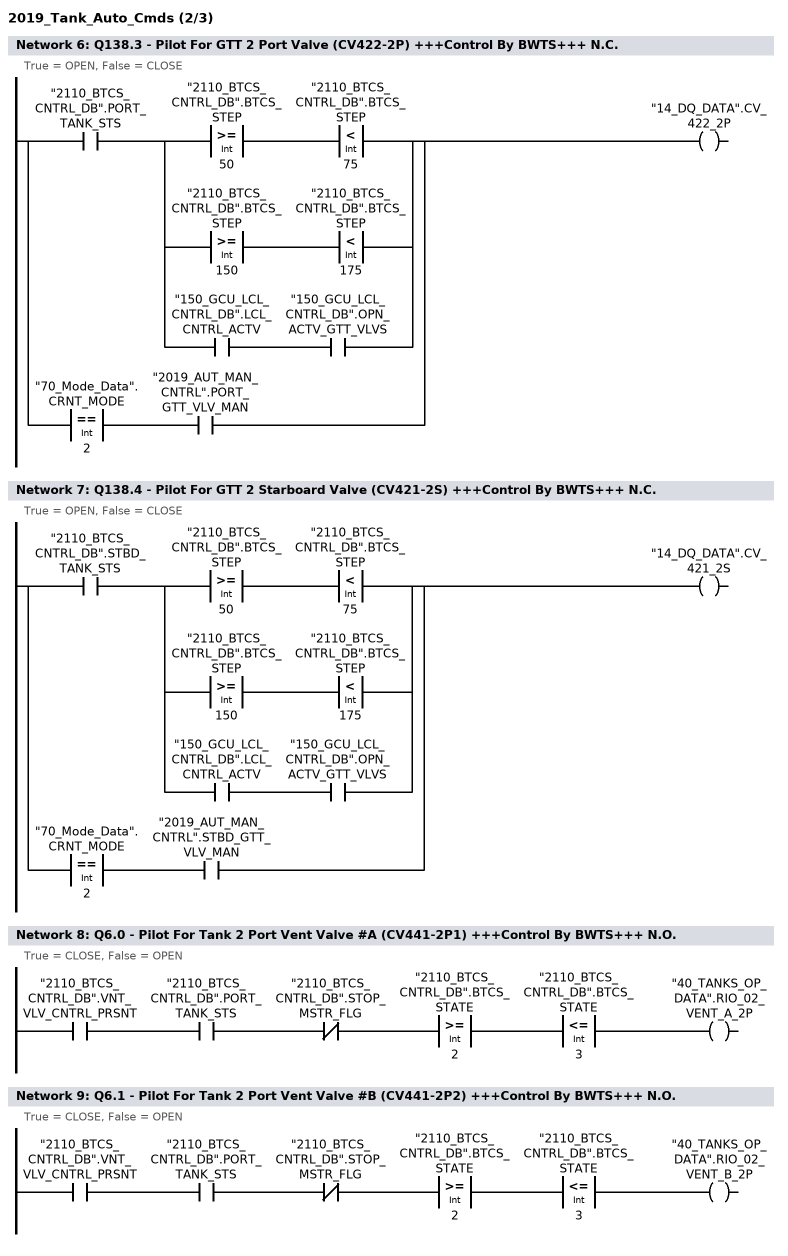
   RUNG wire#powerrail
      Contact( "2110_BTCS_CNTRL_DB".PORT_TANK_STS )
      wire#w1
      { S7_Templates := "SrcType := Int" } GE_Contact(in1 := "2110_BTCS_CNTRL_DB".BTCS_STEP, in2 := 50)
      { S7_Templates := "SrcType := Int" } LT_Contact(in1 := "2110_BTCS_CNTRL_DB".BTCS_STEP, in2 := 75)
      wire#w2
      Coil( "14_DQ_DATA".CV_422_2P )
   END_RUNG
   RUNG wire#w1
      { S7_Templates := "SrcType := Int" } GE_Contact(in1 := "2110_BTCS_CNTRL_DB".BTCS_STEP, in2 := 150)
      { S7_Templates := "SrcType := Int" } LT_Contact(in1 := "2110_BTCS_CNTRL_DB".BTCS_STEP, in2 := 175)
   END_RUNG wire#w2
   RUNG wire#w1
      Contact( "150_GCU_LCL_CNTRL_DB".LCL_CNTRL_ACTV )
      Contact( "150_GCU_LCL_CNTRL_DB".OPN_ACTV_GTT_VLVS )
   END_RUNG wire#w2
   RUNG wire#powerrail
      { S7_Templates := "SrcType := Int" } EQ_Contact(in1 := "70_Mode_Data".CRNT_MODE, in2 := 2)
      Contact( "2019_AUT_MAN_CNTRL".PORT_GTT_VLV_MAN )
   END_RUNG wire#w2
   // the same network as SCL:
   "14_DQ_DATA".CV_422_2P := ("2110_BTCS_CNTRL_DB".PORT_TANK_STS AND ((("2110_BTCS_CNTRL_DB".BTCS_STEP >= 50) AND ("2110_BTCS_CNTRL_DB".BTCS_STEP < 75)) OR (("2110_BTCS_CNTRL_DB".BTCS_STEP >= 150) AND ("2110_BTCS_CNTRL_DB".BTCS_STEP < 175)) OR ("150_GCU_LCL_CNTRL_DB".LCL_CNTRL_ACTV AND "150_GCU_LCL_CNTRL_DB".OPN_ACTV_GTT_VLVS))) OR (("70_Mode_Data".CRNT_MODE = 2) AND "2019_AUT_MAN_CNTRL".PORT_GTT_VLV_MAN);
END_REGION

REGION Network 7: Q138.4 - Pilot For GTT 2 Starboard Valve (CV421-2S) +++Control By BWTS+++ N.C.
   // True = OPEN, False = CLOSE
   RUNG wire#powerrail
      Contact( "2110_BTCS_CNTRL_DB".STBD_TANK_STS )
      wire#w1
      { S7_Templates := "SrcType := Int" } GE_Contact(in1 := "2110_BTCS_CNTRL_DB".BTCS_STEP, in2 := 50)
      { S7_Templates := "SrcType := Int" } LT_Contact(in1 := "2110_BTCS_CNTRL_DB".BTCS_STEP, in2 := 75)
      wire#w2
      Coil( "14_DQ_DATA".CV_421_2S )
   END_RUNG
   RUNG wire#w1
      { S7_Templates := "SrcType := Int" } GE_Contact(in1 := "2110_BTCS_CNTRL_DB".BTCS_STEP, in2 := 150)
      { S7_Templates := "SrcType := Int" } LT_Contact(in1 := "2110_BTCS_CNTRL_DB".BTCS_STEP, in2 := 175)
   END_RUNG wire#w2
   RUNG wire#w1
      Contact( "150_GCU_LCL_CNTRL_DB".LCL_CNTRL_ACTV )
      Contact( "150_GCU_LCL_CNTRL_DB".OPN_ACTV_GTT_VLVS )
   END_RUNG wire#w2
   RUNG wire#powerrail
      { S7_Templates := "SrcType := Int" } EQ_Contact(in1 := "70_Mode_Data".CRNT_MODE, in2 := 2)
      Contact( "2019_AUT_MAN_CNTRL".STBD_GTT_VLV_MAN )
   END_RUNG wire#w2
   // the same network as SCL:
   "14_DQ_DATA".CV_421_2S := ("2110_BTCS_CNTRL_DB".STBD_TANK_STS AND ((("2110_BTCS_CNTRL_DB".BTCS_STEP >= 50) AND ("2110_BTCS_CNTRL_DB".BTCS_STEP < 75)) OR (("2110_BTCS_CNTRL_DB".BTCS_STEP >= 150) AND ("2110_BTCS_CNTRL_DB".BTCS_STEP < 175)) OR ("150_GCU_LCL_CNTRL_DB".LCL_CNTRL_ACTV AND "150_GCU_LCL_CNTRL_DB".OPN_ACTV_GTT_VLVS))) OR (("70_Mode_Data".CRNT_MODE = 2) AND "2019_AUT_MAN_CNTRL".STBD_GTT_VLV_MAN);
END_REGION

REGION Network 8: Q6.0 - Pilot For Tank 2 Port Vent Valve #A (CV441-2P1) +++Control By BWTS+++ N.O.
   // True = CLOSE, False = OPEN
   RUNG wire#powerrail
      Contact( "2110_BTCS_CNTRL_DB".VNT_VLV_CNTRL_PRSNT )
      Contact( "2110_BTCS_CNTRL_DB".PORT_TANK_STS )
      I_Contact( "2110_BTCS_CNTRL_DB".STOP_MSTR_FLG )
      { S7_Templates := "SrcType := Int" } GE_Contact(in1 := "2110_BTCS_CNTRL_DB".BTCS_STATE, in2 := 2)
      { S7_Templates := "SrcType := Int" } LE_Contact(in1 := "2110_BTCS_CNTRL_DB".BTCS_STATE, in2 := 3)
      Coil( "40_TANKS_OP_DATA".RIO_02_VENT_A_2P )
   END_RUNG
   // the same network as SCL:
   "40_TANKS_OP_DATA".RIO_02_VENT_A_2P := "2110_BTCS_CNTRL_DB".VNT_VLV_CNTRL_PRSNT AND "2110_BTCS_CNTRL_DB".PORT_TANK_STS AND NOT "2110_BTCS_CNTRL_DB".STOP_MSTR_FLG AND ("2110_BTCS_CNTRL_DB".BTCS_STATE >= 2) AND ("2110_BTCS_CNTRL_DB".BTCS_STATE <= 3);
END_REGION

REGION Network 9: Q6.1 - Pilot For Tank 2 Port Vent Valve #B (CV441-2P2) +++Control By BWTS+++ N.O.
   // True = CLOSE, False = OPEN
   RUNG wire#powerrail
      Contact( "2110_BTCS_CNTRL_DB".VNT_VLV_CNTRL_PRSNT )
      Contact( "2110_BTCS_CNTRL_DB".PORT_TANK_STS )
      I_Contact( "2110_BTCS_CNTRL_DB".STOP_MSTR_FLG )
      { S7_Templates := "SrcType := Int" } GE_Contact(in1 := "2110_BTCS_CNTRL_DB".BTCS_STATE, in2 := 2)
      { S7_Templates := "SrcType := Int" } LE_Contact(in1 := "2110_BTCS_CNTRL_DB".BTCS_STATE, in2 := 3)
      Coil( "40_TANKS_OP_DATA".RIO_02_VENT_B_2P )
   END_RUNG
   // the same network as SCL:
   "40_TANKS_OP_DATA".RIO_02_VENT_B_2P := "2110_BTCS_CNTRL_DB".VNT_VLV_CNTRL_PRSNT AND "2110_BTCS_CNTRL_DB".PORT_TANK_STS AND NOT "2110_BTCS_CNTRL_DB".STOP_MSTR_FLG AND ("2110_BTCS_CNTRL_DB".BTCS_STATE >= 2) AND ("2110_BTCS_CNTRL_DB".BTCS_STATE <= 3);
END_REGION

REGION Network 10: Q6.2 - Pilot For Tank 2 Starboard Vent Valve #A (CV440-2P1) +++Control By BWTS+++ N.O.
   // True = CLOSE, False = OPEN
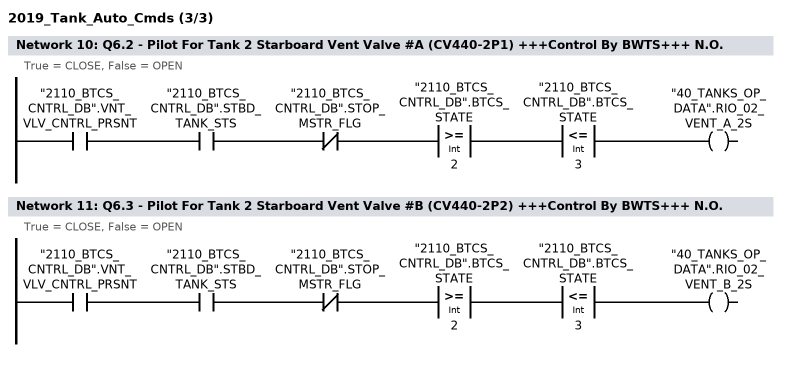
   RUNG wire#powerrail
      Contact( "2110_BTCS_CNTRL_DB".VNT_VLV_CNTRL_PRSNT )
      Contact( "2110_BTCS_CNTRL_DB".STBD_TANK_STS )
      I_Contact( "2110_BTCS_CNTRL_DB".STOP_MSTR_FLG )
      { S7_Templates := "SrcType := Int" } GE_Contact(in1 := "2110_BTCS_CNTRL_DB".BTCS_STATE, in2 := 2)
      { S7_Templates := "SrcType := Int" } LE_Contact(in1 := "2110_BTCS_CNTRL_DB".BTCS_STATE, in2 := 3)
      Coil( "40_TANKS_OP_DATA".RIO_02_VENT_A_2S )
   END_RUNG
   // the same network as SCL:
   "40_TANKS_OP_DATA".RIO_02_VENT_A_2S := "2110_BTCS_CNTRL_DB".VNT_VLV_CNTRL_PRSNT AND "2110_BTCS_CNTRL_DB".STBD_TANK_STS AND NOT "2110_BTCS_CNTRL_DB".STOP_MSTR_FLG AND ("2110_BTCS_CNTRL_DB".BTCS_STATE >= 2) AND ("2110_BTCS_CNTRL_DB".BTCS_STATE <= 3);
END_REGION

REGION Network 11: Q6.3 - Pilot For Tank 2 Starboard Vent Valve #B (CV440-2P2) +++Control By BWTS+++ N.O.
   // True = CLOSE, False = OPEN
   RUNG wire#powerrail
      Contact( "2110_BTCS_CNTRL_DB".VNT_VLV_CNTRL_PRSNT )
      Contact( "2110_BTCS_CNTRL_DB".STBD_TANK_STS )
      I_Contact( "2110_BTCS_CNTRL_DB".STOP_MSTR_FLG )
      { S7_Templates := "SrcType := Int" } GE_Contact(in1 := "2110_BTCS_CNTRL_DB".BTCS_STATE, in2 := 2)
      { S7_Templates := "SrcType := Int" } LE_Contact(in1 := "2110_BTCS_CNTRL_DB".BTCS_STATE, in2 := 3)
      Coil( "40_TANKS_OP_DATA".RIO_02_VENT_B_2S )
   END_RUNG
   // the same network as SCL:
   "40_TANKS_OP_DATA".RIO_02_VENT_B_2S := "2110_BTCS_CNTRL_DB".VNT_VLV_CNTRL_PRSNT AND "2110_BTCS_CNTRL_DB".STBD_TANK_STS AND NOT "2110_BTCS_CNTRL_DB".STOP_MSTR_FLG AND ("2110_BTCS_CNTRL_DB".BTCS_STATE >= 2) AND ("2110_BTCS_CNTRL_DB".BTCS_STATE <= 3);
END_REGION
END_FUNCTION_BLOCK

FUNCTION "2019_AUTO_CMNDS" : Void   // FC2019, LAD
TITLE = Automatic Output Commands
{ S7_Optimized_Access := 'TRUE' }
AUTHOR : JRS
VERSION : 0.1
// To process automatic output commands prior to output processing
BEGIN

REGION Network 1: Q136.2 - Block Valve 1 Control (CV407) +++Control By BWTS+++ N.C.
   // True = OPEN, False = CLOSE
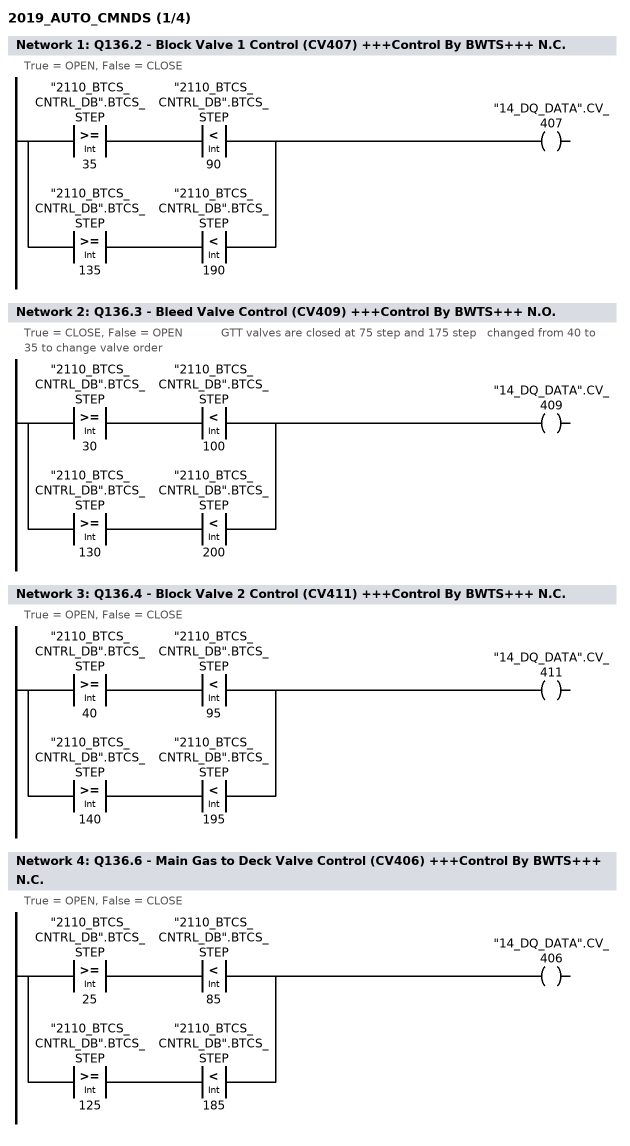
   RUNG wire#powerrail
      { S7_Templates := "SrcType := Int" } GE_Contact(in1 := "2110_BTCS_CNTRL_DB".BTCS_STEP, in2 := 35)
      { S7_Templates := "SrcType := Int" } LT_Contact(in1 := "2110_BTCS_CNTRL_DB".BTCS_STEP, in2 := 90)
      wire#w1
      Coil( "14_DQ_DATA".CV_407 )
   END_RUNG
   RUNG wire#powerrail
      { S7_Templates := "SrcType := Int" } GE_Contact(in1 := "2110_BTCS_CNTRL_DB".BTCS_STEP, in2 := 135)
      { S7_Templates := "SrcType := Int" } LT_Contact(in1 := "2110_BTCS_CNTRL_DB".BTCS_STEP, in2 := 190)
   END_RUNG wire#w1
   // the same network as SCL:
   "14_DQ_DATA".CV_407 := (("2110_BTCS_CNTRL_DB".BTCS_STEP >= 35) AND ("2110_BTCS_CNTRL_DB".BTCS_STEP < 90)) OR (("2110_BTCS_CNTRL_DB".BTCS_STEP >= 135) AND ("2110_BTCS_CNTRL_DB".BTCS_STEP < 190));
END_REGION

REGION Network 2: Q136.3 - Bleed Valve Control (CV409) +++Control By BWTS+++ N.O.
   // True = CLOSE, False = OPEN           GTT valves are closed at 75 step and 175 step   changed from 40 to 35 to change valve order
   RUNG wire#powerrail
      { S7_Templates := "SrcType := Int" } GE_Contact(in1 := "2110_BTCS_CNTRL_DB".BTCS_STEP, in2 := 30)
      { S7_Templates := "SrcType := Int" } LT_Contact(in1 := "2110_BTCS_CNTRL_DB".BTCS_STEP, in2 := 100)
      wire#w1
      Coil( "14_DQ_DATA".CV_409 )
   END_RUNG
   RUNG wire#powerrail
      { S7_Templates := "SrcType := Int" } GE_Contact(in1 := "2110_BTCS_CNTRL_DB".BTCS_STEP, in2 := 130)
      { S7_Templates := "SrcType := Int" } LT_Contact(in1 := "2110_BTCS_CNTRL_DB".BTCS_STEP, in2 := 200)
   END_RUNG wire#w1
   // the same network as SCL:
   "14_DQ_DATA".CV_409 := (("2110_BTCS_CNTRL_DB".BTCS_STEP >= 30) AND ("2110_BTCS_CNTRL_DB".BTCS_STEP < 100)) OR (("2110_BTCS_CNTRL_DB".BTCS_STEP >= 130) AND ("2110_BTCS_CNTRL_DB".BTCS_STEP < 200));
END_REGION

REGION Network 3: Q136.4 - Block Valve 2 Control (CV411) +++Control By BWTS+++ N.C.
   // True = OPEN, False = CLOSE
   RUNG wire#powerrail
      { S7_Templates := "SrcType := Int" } GE_Contact(in1 := "2110_BTCS_CNTRL_DB".BTCS_STEP, in2 := 40)
      { S7_Templates := "SrcType := Int" } LT_Contact(in1 := "2110_BTCS_CNTRL_DB".BTCS_STEP, in2 := 95)
      wire#w1
      Coil( "14_DQ_DATA".CV_411 )
   END_RUNG
   RUNG wire#powerrail
      { S7_Templates := "SrcType := Int" } GE_Contact(in1 := "2110_BTCS_CNTRL_DB".BTCS_STEP, in2 := 140)
      { S7_Templates := "SrcType := Int" } LT_Contact(in1 := "2110_BTCS_CNTRL_DB".BTCS_STEP, in2 := 195)
   END_RUNG wire#w1
   // the same network as SCL:
   "14_DQ_DATA".CV_411 := (("2110_BTCS_CNTRL_DB".BTCS_STEP >= 40) AND ("2110_BTCS_CNTRL_DB".BTCS_STEP < 95)) OR (("2110_BTCS_CNTRL_DB".BTCS_STEP >= 140) AND ("2110_BTCS_CNTRL_DB".BTCS_STEP < 195));
END_REGION

REGION Network 4: Q136.6 - Main Gas to Deck Valve Control (CV406) +++Control By BWTS+++ N.C.
   // True = OPEN, False = CLOSE
   RUNG wire#powerrail
      { S7_Templates := "SrcType := Int" } GE_Contact(in1 := "2110_BTCS_CNTRL_DB".BTCS_STEP, in2 := 25)
      { S7_Templates := "SrcType := Int" } LT_Contact(in1 := "2110_BTCS_CNTRL_DB".BTCS_STEP, in2 := 85)
      wire#w1
      Coil( "14_DQ_DATA".CV_406 )
   END_RUNG
   RUNG wire#powerrail
      { S7_Templates := "SrcType := Int" } GE_Contact(in1 := "2110_BTCS_CNTRL_DB".BTCS_STEP, in2 := 125)
      { S7_Templates := "SrcType := Int" } LT_Contact(in1 := "2110_BTCS_CNTRL_DB".BTCS_STEP, in2 := 185)
   END_RUNG wire#w1
   // the same network as SCL:
   "14_DQ_DATA".CV_406 := (("2110_BTCS_CNTRL_DB".BTCS_STEP >= 25) AND ("2110_BTCS_CNTRL_DB".BTCS_STEP < 85)) OR (("2110_BTCS_CNTRL_DB".BTCS_STEP >= 125) AND ("2110_BTCS_CNTRL_DB".BTCS_STEP < 185));
END_REGION

REGION Network 5: TANK TREATMENT RUN DE-OX/RE-OX -(Q138.3 - Pilot For GTT 2 Port Valve (CV422-2P) +++Control By BWTS+++ N.C.)
   // True = OPEN, False = CLOSE
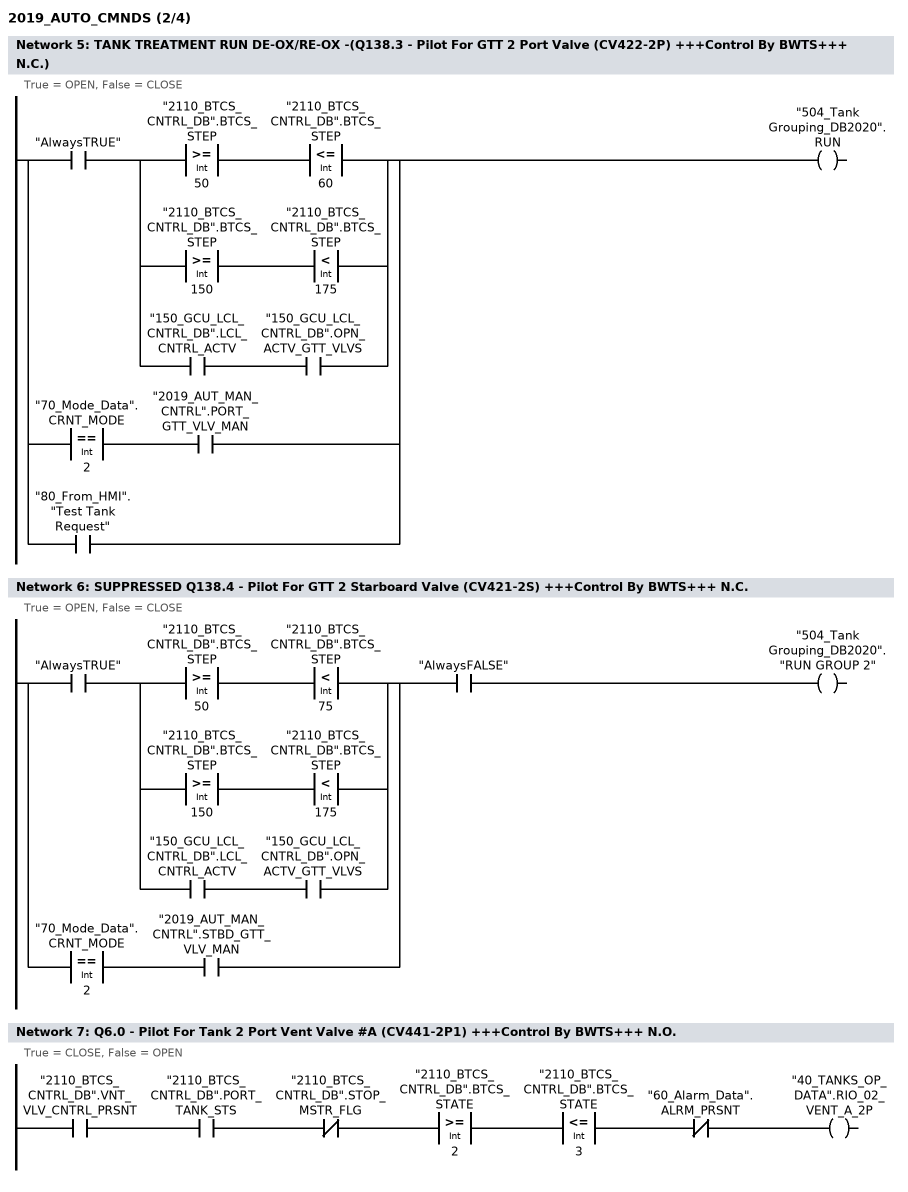
   RUNG wire#powerrail
      Contact( "AlwaysTRUE" )
      wire#w1
      { S7_Templates := "SrcType := Int" } GE_Contact(in1 := "2110_BTCS_CNTRL_DB".BTCS_STEP, in2 := 50)
      { S7_Templates := "SrcType := Int" } LE_Contact(in1 := "2110_BTCS_CNTRL_DB".BTCS_STEP, in2 := 60)
      wire#w2
      Coil( "504_Tank Grouping_DB2020".RUN )
   END_RUNG
   RUNG wire#w1
      { S7_Templates := "SrcType := Int" } GE_Contact(in1 := "2110_BTCS_CNTRL_DB".BTCS_STEP, in2 := 150)
      { S7_Templates := "SrcType := Int" } LT_Contact(in1 := "2110_BTCS_CNTRL_DB".BTCS_STEP, in2 := 175)
   END_RUNG wire#w2
   RUNG wire#w1
      Contact( "150_GCU_LCL_CNTRL_DB".LCL_CNTRL_ACTV )
      Contact( "150_GCU_LCL_CNTRL_DB".OPN_ACTV_GTT_VLVS )
   END_RUNG wire#w2
   RUNG wire#powerrail
      { S7_Templates := "SrcType := Int" } EQ_Contact(in1 := "70_Mode_Data".CRNT_MODE, in2 := 2)
      Contact( "2019_AUT_MAN_CNTRL".PORT_GTT_VLV_MAN )
   END_RUNG wire#w2
   RUNG wire#powerrail
      Contact( "80_From_HMI"."Test Tank Request" )
   END_RUNG wire#w2
   // the same network as SCL:
   "504_Tank Grouping_DB2020".RUN := ("AlwaysTRUE" AND ((("2110_BTCS_CNTRL_DB".BTCS_STEP >= 50) AND ("2110_BTCS_CNTRL_DB".BTCS_STEP <= 60)) OR (("2110_BTCS_CNTRL_DB".BTCS_STEP >= 150) AND ("2110_BTCS_CNTRL_DB".BTCS_STEP < 175)) OR ("150_GCU_LCL_CNTRL_DB".LCL_CNTRL_ACTV AND "150_GCU_LCL_CNTRL_DB".OPN_ACTV_GTT_VLVS))) OR (("70_Mode_Data".CRNT_MODE = 2) AND "2019_AUT_MAN_CNTRL".PORT_GTT_VLV_MAN) OR "80_From_HMI"."Test Tank Request";
END_REGION

REGION Network 6: SUPPRESSED Q138.4 - Pilot For GTT 2 Starboard Valve (CV421-2S) +++Control By BWTS+++ N.C.
   // True = OPEN, False = CLOSE
   RUNG wire#powerrail
      Contact( "AlwaysTRUE" )
      wire#w1
      { S7_Templates := "SrcType := Int" } GE_Contact(in1 := "2110_BTCS_CNTRL_DB".BTCS_STEP, in2 := 50)
      { S7_Templates := "SrcType := Int" } LT_Contact(in1 := "2110_BTCS_CNTRL_DB".BTCS_STEP, in2 := 75)
      wire#w2
      Contact( "AlwaysFALSE" )
      Coil( "504_Tank Grouping_DB2020"."RUN GROUP 2" )
   END_RUNG
   RUNG wire#w1
      { S7_Templates := "SrcType := Int" } GE_Contact(in1 := "2110_BTCS_CNTRL_DB".BTCS_STEP, in2 := 150)
      { S7_Templates := "SrcType := Int" } LT_Contact(in1 := "2110_BTCS_CNTRL_DB".BTCS_STEP, in2 := 175)
   END_RUNG wire#w2
   RUNG wire#w1
      Contact( "150_GCU_LCL_CNTRL_DB".LCL_CNTRL_ACTV )
      Contact( "150_GCU_LCL_CNTRL_DB".OPN_ACTV_GTT_VLVS )
   END_RUNG wire#w2
   RUNG wire#powerrail
      { S7_Templates := "SrcType := Int" } EQ_Contact(in1 := "70_Mode_Data".CRNT_MODE, in2 := 2)
      Contact( "2019_AUT_MAN_CNTRL".STBD_GTT_VLV_MAN )
   END_RUNG wire#w2
   // the same network as SCL:
   "504_Tank Grouping_DB2020"."RUN GROUP 2" := (("AlwaysTRUE" AND ((("2110_BTCS_CNTRL_DB".BTCS_STEP >= 50) AND ("2110_BTCS_CNTRL_DB".BTCS_STEP < 75)) OR (("2110_BTCS_CNTRL_DB".BTCS_STEP >= 150) AND ("2110_BTCS_CNTRL_DB".BTCS_STEP < 175)) OR ("150_GCU_LCL_CNTRL_DB".LCL_CNTRL_ACTV AND "150_GCU_LCL_CNTRL_DB".OPN_ACTV_GTT_VLVS))) OR (("70_Mode_Data".CRNT_MODE = 2) AND "2019_AUT_MAN_CNTRL".STBD_GTT_VLV_MAN)) AND "AlwaysFALSE";
END_REGION

REGION Network 7: Q6.0 - Pilot For Tank 2 Port Vent Valve #A (CV441-2P1) +++Control By BWTS+++ N.O.
   // True = CLOSE, False = OPEN
   RUNG wire#powerrail
      Contact( "2110_BTCS_CNTRL_DB".VNT_VLV_CNTRL_PRSNT )
      Contact( "2110_BTCS_CNTRL_DB".PORT_TANK_STS )
      I_Contact( "2110_BTCS_CNTRL_DB".STOP_MSTR_FLG )
      { S7_Templates := "SrcType := Int" } GE_Contact(in1 := "2110_BTCS_CNTRL_DB".BTCS_STATE, in2 := 2)
      { S7_Templates := "SrcType := Int" } LE_Contact(in1 := "2110_BTCS_CNTRL_DB".BTCS_STATE, in2 := 3)
      I_Contact( "60_Alarm_Data".ALRM_PRSNT )
      Coil( "40_TANKS_OP_DATA".RIO_02_VENT_A_2P )
   END_RUNG
   // the same network as SCL:
   "40_TANKS_OP_DATA".RIO_02_VENT_A_2P := "2110_BTCS_CNTRL_DB".VNT_VLV_CNTRL_PRSNT AND "2110_BTCS_CNTRL_DB".PORT_TANK_STS AND NOT "2110_BTCS_CNTRL_DB".STOP_MSTR_FLG AND ("2110_BTCS_CNTRL_DB".BTCS_STATE >= 2) AND ("2110_BTCS_CNTRL_DB".BTCS_STATE <= 3) AND NOT "60_Alarm_Data".ALRM_PRSNT;
END_REGION

REGION Network 8: Q6.1 - Pilot For Tank 2 Port Vent Valve #B (CV441-2P2) +++Control By BWTS+++ N.O.
   // True = CLOSE, False = OPEN
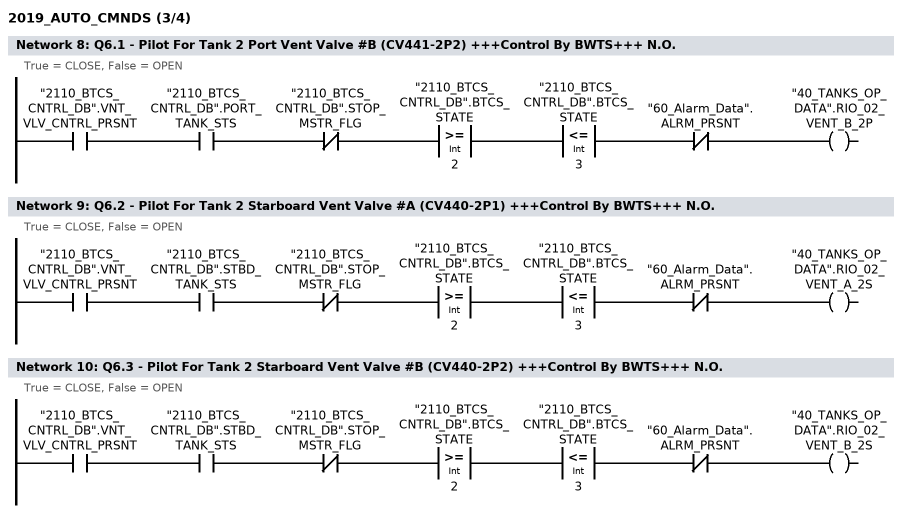
   RUNG wire#powerrail
      Contact( "2110_BTCS_CNTRL_DB".VNT_VLV_CNTRL_PRSNT )
      Contact( "2110_BTCS_CNTRL_DB".PORT_TANK_STS )
      I_Contact( "2110_BTCS_CNTRL_DB".STOP_MSTR_FLG )
      { S7_Templates := "SrcType := Int" } GE_Contact(in1 := "2110_BTCS_CNTRL_DB".BTCS_STATE, in2 := 2)
      { S7_Templates := "SrcType := Int" } LE_Contact(in1 := "2110_BTCS_CNTRL_DB".BTCS_STATE, in2 := 3)
      I_Contact( "60_Alarm_Data".ALRM_PRSNT )
      Coil( "40_TANKS_OP_DATA".RIO_02_VENT_B_2P )
   END_RUNG
   // the same network as SCL:
   "40_TANKS_OP_DATA".RIO_02_VENT_B_2P := "2110_BTCS_CNTRL_DB".VNT_VLV_CNTRL_PRSNT AND "2110_BTCS_CNTRL_DB".PORT_TANK_STS AND NOT "2110_BTCS_CNTRL_DB".STOP_MSTR_FLG AND ("2110_BTCS_CNTRL_DB".BTCS_STATE >= 2) AND ("2110_BTCS_CNTRL_DB".BTCS_STATE <= 3) AND NOT "60_Alarm_Data".ALRM_PRSNT;
END_REGION

REGION Network 9: Q6.2 - Pilot For Tank 2 Starboard Vent Valve #A (CV440-2P1) +++Control By BWTS+++ N.O.
   // True = CLOSE, False = OPEN
   RUNG wire#powerrail
      Contact( "2110_BTCS_CNTRL_DB".VNT_VLV_CNTRL_PRSNT )
      Contact( "2110_BTCS_CNTRL_DB".STBD_TANK_STS )
      I_Contact( "2110_BTCS_CNTRL_DB".STOP_MSTR_FLG )
      { S7_Templates := "SrcType := Int" } GE_Contact(in1 := "2110_BTCS_CNTRL_DB".BTCS_STATE, in2 := 2)
      { S7_Templates := "SrcType := Int" } LE_Contact(in1 := "2110_BTCS_CNTRL_DB".BTCS_STATE, in2 := 3)
      I_Contact( "60_Alarm_Data".ALRM_PRSNT )
      Coil( "40_TANKS_OP_DATA".RIO_02_VENT_A_2S )
   END_RUNG
   // the same network as SCL:
   "40_TANKS_OP_DATA".RIO_02_VENT_A_2S := "2110_BTCS_CNTRL_DB".VNT_VLV_CNTRL_PRSNT AND "2110_BTCS_CNTRL_DB".STBD_TANK_STS AND NOT "2110_BTCS_CNTRL_DB".STOP_MSTR_FLG AND ("2110_BTCS_CNTRL_DB".BTCS_STATE >= 2) AND ("2110_BTCS_CNTRL_DB".BTCS_STATE <= 3) AND NOT "60_Alarm_Data".ALRM_PRSNT;
END_REGION

REGION Network 10: Q6.3 - Pilot For Tank 2 Starboard Vent Valve #B (CV440-2P2) +++Control By BWTS+++ N.O.
   // True = CLOSE, False = OPEN
   RUNG wire#powerrail
      Contact( "2110_BTCS_CNTRL_DB".VNT_VLV_CNTRL_PRSNT )
      Contact( "2110_BTCS_CNTRL_DB".STBD_TANK_STS )
      I_Contact( "2110_BTCS_CNTRL_DB".STOP_MSTR_FLG )
      { S7_Templates := "SrcType := Int" } GE_Contact(in1 := "2110_BTCS_CNTRL_DB".BTCS_STATE, in2 := 2)
      { S7_Templates := "SrcType := Int" } LE_Contact(in1 := "2110_BTCS_CNTRL_DB".BTCS_STATE, in2 := 3)
      I_Contact( "60_Alarm_Data".ALRM_PRSNT )
      Coil( "40_TANKS_OP_DATA".RIO_02_VENT_B_2S )
   END_RUNG
   // the same network as SCL:
   "40_TANKS_OP_DATA".RIO_02_VENT_B_2S := "2110_BTCS_CNTRL_DB".VNT_VLV_CNTRL_PRSNT AND "2110_BTCS_CNTRL_DB".STBD_TANK_STS AND NOT "2110_BTCS_CNTRL_DB".STOP_MSTR_FLG AND ("2110_BTCS_CNTRL_DB".BTCS_STATE >= 2) AND ("2110_BTCS_CNTRL_DB".BTCS_STATE <= 3) AND NOT "60_Alarm_Data".ALRM_PRSNT;
END_REGION

REGION Network 11: Tank Grouping
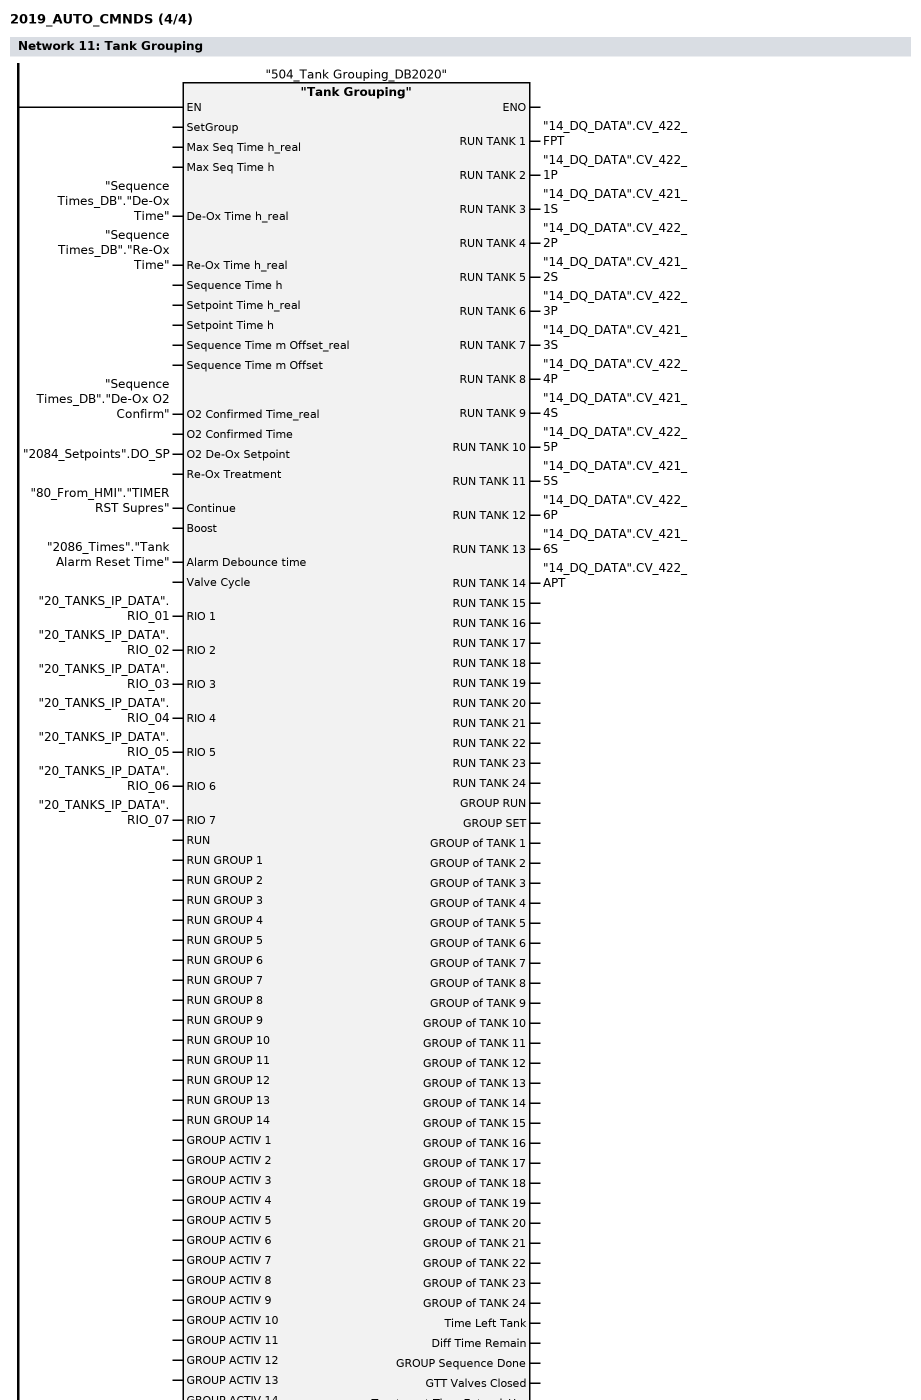
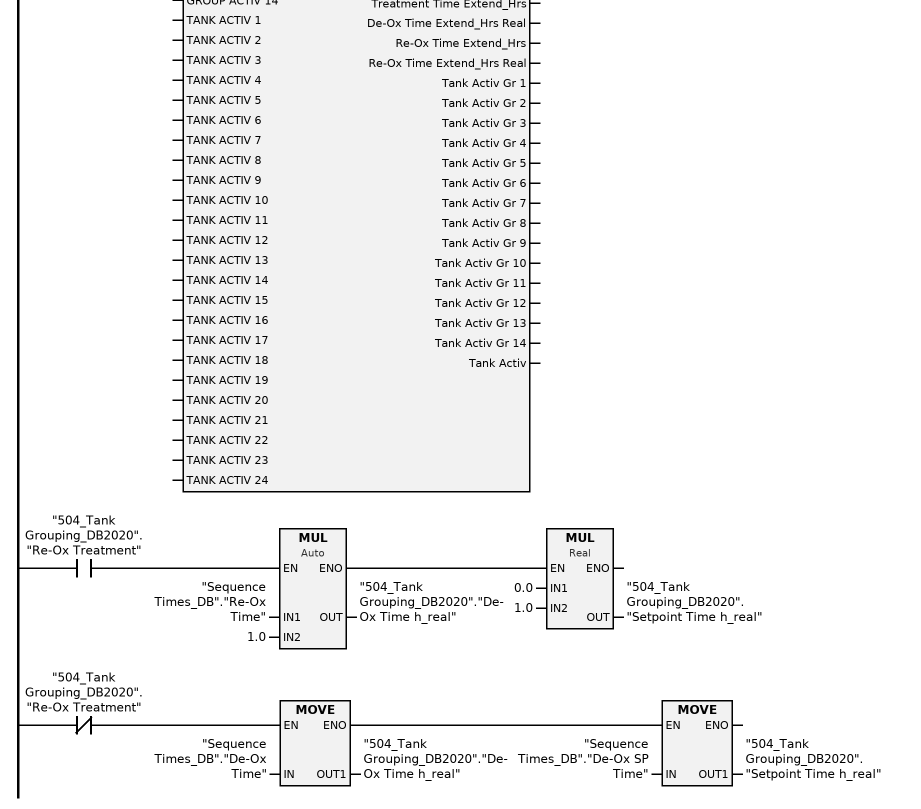
   RUNG wire#powerrail
      "504_Tank Grouping_DB2020"(SetGroup :=, "Max Seq Time h_real" :=, "Max Seq Time h" :=, "De-Ox Time h_real" := "Sequence Times_DB"."De-Ox Time", "Re-Ox Time h_real" := "Sequence Times_DB"."Re-Ox Time", "Sequence Time h" :=, "Setpoint Time h_real" :=, "Setpoint Time h" :=, "Sequence Time m Offset_real" :=, "Sequence Time m Offset" :=, "O2 Confirmed Time_real" := "Sequence Times_DB"."De-Ox O2 Confirm", "O2 Confirmed Time" :=, "O2 De-Ox Setpoint" := "2084_Setpoints".DO_SP, "Re-Ox Treatment" :=, Continue := "80_From_HMI"."TIMER RST Supres", Boost :=, "Alarm Debounce time" := "2086_Times"."Tank Alarm Reset Time", "Valve Cycle" :=, "RIO 1" := "20_TANKS_IP_DATA".RIO_01, "RIO 2" := "20_TANKS_IP_DATA".RIO_02, "RIO 3" := "20_TANKS_IP_DATA".RIO_03, "RIO 4" := "20_TANKS_IP_DATA".RIO_04, "RIO 5" := "20_TANKS_IP_DATA".RIO_05, "RIO 6" := "20_TANKS_IP_DATA".RIO_06, "RIO 7" := "20_TANKS_IP_DATA".RIO_07, RUN :=, "RUN GROUP 1" :=, "RUN GROUP 2" :=, "RUN GROUP 3" :=, "RUN GROUP 4" :=, "RUN GROUP 5" :=, "RUN GROUP 6" :=, "RUN GROUP 7" :=, "RUN GROUP 8" :=, "RUN GROUP 9" :=, "RUN GROUP 10" :=, "RUN GROUP 11" :=, "RUN GROUP 12" :=, "RUN GROUP 13" :=, "RUN GROUP 14" :=, "GROUP ACTIV 1" :=, "GROUP ACTIV 2" :=, "GROUP ACTIV 3" :=, "GROUP ACTIV 4" :=, "GROUP ACTIV 5" :=, "GROUP ACTIV 6" :=, "GROUP ACTIV 7" :=, "GROUP ACTIV 8" :=, "GROUP ACTIV 9" :=, "GROUP ACTIV 10" :=, "GROUP ACTIV 11" :=, "GROUP ACTIV 12" :=, "GROUP ACTIV 13" :=, "GROUP ACTIV 14" :=, "TANK ACTIV 1" :=, "TANK ACTIV 2" :=, "TANK ACTIV 3" :=, "TANK ACTIV 4" :=, "TANK ACTIV 5" :=, "TANK ACTIV 6" :=, "TANK ACTIV 7" :=, "TANK ACTIV 8" :=, "TANK ACTIV 9" :=, "TANK ACTIV 10" :=, "TANK ACTIV 11" :=, "TANK ACTIV 12" :=, "TANK ACTIV 13" :=, "TANK ACTIV 14" :=, "TANK ACTIV 15" :=, "TANK ACTIV 16" :=, "TANK ACTIV 17" :=, "TANK ACTIV 18" :=, "TANK ACTIV 19" :=, "TANK ACTIV 20" :=, "TANK ACTIV 21" :=, "TANK ACTIV 22" :=, "TANK ACTIV 23" :=, "TANK ACTIV 24" :=, "RUN TANK 1" => "14_DQ_DATA".CV_422_FPT, "RUN TANK 2" => "14_DQ_DATA".CV_422_1P, "RUN TANK 3" => "14_DQ_DATA".CV_421_1S, "RUN TANK 4" => "14_DQ_DATA".CV_422_2P, "RUN TANK 5" => "14_DQ_DATA".CV_421_2S, "RUN TANK 6" => "14_DQ_DATA".CV_422_3P, "RUN TANK 7" => "14_DQ_DATA".CV_421_3S, "RUN TANK 8" => "14_DQ_DATA".CV_422_4P, "RUN TANK 9" => "14_DQ_DATA".CV_421_4S, "RUN TANK 10" => "14_DQ_DATA".CV_422_5P, "RUN TANK 11" => "14_DQ_DATA".CV_421_5S, "RUN TANK 12" => "14_DQ_DATA".CV_422_6P, "RUN TANK 13" => "14_DQ_DATA".CV_421_6S, "RUN TANK 14" => "14_DQ_DATA".CV_422_APT, "RUN TANK 15" =>, "RUN TANK 16" =>, "RUN TANK 17" =>, "RUN TANK 18" =>, "RUN TANK 19" =>, "RUN TANK 20" =>, "RUN TANK 21" =>, "RUN TANK 22" =>, "RUN TANK 23" =>, "RUN TANK 24" =>, "GROUP RUN" =>, "GROUP SET" =>, "GROUP of TANK 1" =>, "GROUP of TANK 2" =>, "GROUP of TANK 3" =>, "GROUP of TANK 4" =>, "GROUP of TANK 5" =>, "GROUP of TANK 6" =>, "GROUP of TANK 7" =>, "GROUP of TANK 8" =>, "GROUP of TANK 9" =>, "GROUP of TANK 10" =>, "GROUP of TANK 11" =>, "GROUP of TANK 12" =>, "GROUP of TANK 13" =>, "GROUP of TANK 14" =>, "GROUP of TANK 15" =>, "GROUP of TANK 16" =>, "GROUP of TANK 17" =>, "GROUP of TANK 18" =>, "GROUP of TANK 19" =>, "GROUP of TANK 20" =>, "GROUP of TANK 21" =>, "GROUP of TANK 22" =>, "GROUP of TANK 23" =>, "GROUP of TANK 24" =>, "Time Left Tank" =>, "Diff Time Remain" =>, "GROUP Sequence Done" =>, "GTT Valves Closed" =>, "Treatment Time Extend_Hrs" =>, "De-Ox Time Extend_Hrs Real" =>, "Re-Ox Time Extend_Hrs" =>, "Re-Ox Time Extend_Hrs Real" =>, "Tank Activ Gr 1" =>, "Tank Activ Gr 2" =>, "Tank Activ Gr 3" =>, "Tank Activ Gr 4" =>, "Tank Activ Gr 5" =>, "Tank Activ Gr 6" =>, "Tank Activ Gr 7" =>, "Tank Activ Gr 8" =>, "Tank Activ Gr 9" =>, "Tank Activ Gr 10" =>, "Tank Activ Gr 11" =>, "Tank Activ Gr 12" =>, "Tank Activ Gr 13" =>, "Tank Activ Gr 14" =>, "Tank Activ" =>)
   END_RUNG
   RUNG wire#powerrail
      Contact( "504_Tank Grouping_DB2020"."Re-Ox Treatment" )
      Mul(in1 := "Sequence Times_DB"."Re-Ox Time", in2 := 1.0, out => "504_Tank Grouping_DB2020"."De-Ox Time h_real")
      { S7_Templates := "SrcType := Real" } Mul(in1 := 0.0, in2 := 1.0, out => "504_Tank Grouping_DB2020"."Setpoint Time h_real")
   END_RUNG
   RUNG wire#powerrail
      I_Contact( "504_Tank Grouping_DB2020"."Re-Ox Treatment" )
      Move(in := "Sequence Times_DB"."De-Ox Time", out1 => "504_Tank Grouping_DB2020"."De-Ox Time h_real")
      Move(in := "Sequence Times_DB"."De-Ox SP Time", out1 => "504_Tank Grouping_DB2020"."Setpoint Time h_real")
   END_RUNG
   // the same network as SCL:
   "504_Tank Grouping_DB2020"("De-Ox Time h_real" := "Sequence Times_DB"."De-Ox Time",   // "Tank Grouping"
                           "Re-Ox Time h_real" := "Sequence Times_DB"."Re-Ox Time",
                           "O2 Confirmed Time_real" := "Sequence Times_DB"."De-Ox O2 Confirm",
                           "O2 De-Ox Setpoint" := "2084_Setpoints".DO_SP,
                           Continue := "80_From_HMI"."TIMER RST Supres",
                           "Alarm Debounce time" := "2086_Times"."Tank Alarm Reset Time",
                           "RIO 1" := "20_TANKS_IP_DATA".RIO_01,
                           "RIO 2" := "20_TANKS_IP_DATA".RIO_02,
                           "RIO 3" := "20_TANKS_IP_DATA".RIO_03,
                           "RIO 4" := "20_TANKS_IP_DATA".RIO_04,
                           "RIO 5" := "20_TANKS_IP_DATA".RIO_05,
                           "RIO 6" := "20_TANKS_IP_DATA".RIO_06,
                           "RIO 7" := "20_TANKS_IP_DATA".RIO_07,
                           "RUN TANK 1" => "14_DQ_DATA".CV_422_FPT,
                           "RUN TANK 2" => "14_DQ_DATA".CV_422_1P,
                           "RUN TANK 3" => "14_DQ_DATA".CV_421_1S,
                           "RUN TANK 4" => "14_DQ_DATA".CV_422_2P,
                           "RUN TANK 5" => "14_DQ_DATA".CV_421_2S,
                           "RUN TANK 6" => "14_DQ_DATA".CV_422_3P,
                           "RUN TANK 7" => "14_DQ_DATA".CV_421_3S,
                           "RUN TANK 8" => "14_DQ_DATA".CV_422_4P,
                           "RUN TANK 9" => "14_DQ_DATA".CV_421_4S,
                           "RUN TANK 10" => "14_DQ_DATA".CV_422_5P,
                           "RUN TANK 11" => "14_DQ_DATA".CV_421_5S,
                           "RUN TANK 12" => "14_DQ_DATA".CV_422_6P,
                           "RUN TANK 13" => "14_DQ_DATA".CV_421_6S,
                           "RUN TANK 14" => "14_DQ_DATA".CV_422_APT);
   IF "504_Tank Grouping_DB2020"."Re-Ox Treatment" THEN
       "504_Tank Grouping_DB2020"."De-Ox Time h_real" := "Sequence Times_DB"."Re-Ox Time" * 1.0;
       "504_Tank Grouping_DB2020"."Setpoint Time h_real" := 0.0 * 1.0;
   END_IF;
   IF NOT "504_Tank Grouping_DB2020"."Re-Ox Treatment" THEN
       "504_Tank Grouping_DB2020"."De-Ox Time h_real" := "Sequence Times_DB"."De-Ox Time";
       "504_Tank Grouping_DB2020"."Setpoint Time h_real" := "Sequence Times_DB"."De-Ox SP Time";
   END_IF;
END_REGION
END_FUNCTION

// folder: 2000 - 2999 BTCS System/2050 - 2059 PLC Communication

FUNCTION "2058_PLC_SIGNALS" : Void   // FC2058, LAD
TITLE = PLC Signals
{ S7_Optimized_Access := 'TRUE' }
AUTHOR : JRS
VERSION : 0.1
// For managing the signals between the BTCS and GCU PLC
BEGIN

REGION Network 1: State